// TIA Portal project "FABRICA DE TAPAS - TRANSPORTE -TUNEL DE ENFRIAMIENTO" (V17)

(* hardware
DEVICE "S7-1500/ET200MP station_1"  S7-1500 station
   slot 0: "Rail_0"  Rack  6ES7 590-1***0-0AA0
   slot 1: "CPU_PRINCIPAL"  CPU 1511-1 PN  6ES7 511-1AK02-0AB0  V2.8
      slot 3: "CPU display_1"  6ES7591-1AA00-0AA0
      slot 32768: "PROFINET interface_1"  X1
         slot 32769: "Port_1"  X1 P1
         slot 32770: "Port_2"  X1 P2
      slot 34817: "Virtual CP interface port_1"  Virtual CP interface port  Virtual CP interface port
DEVICE "HMI-TRANSPORTE"  KTP700 Basic PN
   slot 0: "HMI-TRANSPORTE"  KTP700 Basic PN  6AV2 123-2GB03-0AX0  17.0.0.0
   slot 1: "HMI_RT_1"  KTP700 Basic PN  6AV2 123-2GB03-0AX0  17.0.0.0
   slot 5: "HMI-TRANSPORTE.IE_CP_1"  PROFINET Interface  17.0.0.0
      slot 1: "PROFINET Interface_1"  PROFINET Interface
         slot 1: "Port_1"  Port
DEVICE "TUNEL-1"  KTP700 Basic PN
   slot 0: "TUNEL-1"  KTP700 Basic PN  6AV2 123-2GB03-0AX0  17.0.0.0
   slot 1: "HMI_RT_2"  KTP700 Basic PN  6AV2 123-2GB03-0AX0  17.0.0.0
   slot 5: "TUNEL-1.IE_CP_1"  PROFINET Interface  17.0.0.0
      slot 1: "PROFINET Interface_1"  PROFINET Interface
         slot 1: "Port_1"  Port
DEVICE "TUNEL-2"  KTP700 Basic PN
   slot 0: "TUNEL-2"  KTP700 Basic PN  6AV2 123-2GB03-0AX0  17.0.0.0
   slot 1: "HMI_RT_3"  KTP700 Basic PN  6AV2 123-2GB03-0AX0  17.0.0.0
   slot 5: "TUNEL-2.IE_CP_1"  PROFINET Interface  17.0.0.0
      slot 1: "PROFINET Interface_1"  PROFINET Interface
         slot 1: "Port_1"  Port
DEVICE "ET 200SP station_1"  ET 200SP-Station
   slot 0: "Rack_0"  Rack  6ES5 710-8MAx1
   slot 0: "TRANSPORTE"  IM 155-6 PN ST  6ES7 155-6AU01-0BN0  V4.2
   slot 1: "DI 16x24VDC ST_1"  DI 16x24VDC ST  6ES7 131-6BH01-0BA0  V0.0
      slot 1: "DI 16x24VDC ST_1"  DI 16x24VDC ST
   slot 2: "DQ 16x24VDC/0.5A ST_1"  DQ 16x24VDC/0.5A ST  6ES7 132-6BH01-0BA0  V0.0
      slot 1: "DQ 16x24VDC/0.5A ST_1"  DQ 16x24VDC/0.5A ST
   slot 3: "Server module_1"  Server module  6ES7 193-6PA00-0AA0  V1.1
      slot 1: "Server module_1"  Server module
   slot 127: "BA 2xRJ45"  BA 2xRJ45  6ES7 193-6AR00-0AA0  V0.0
      slot 1: "Port_1"  X1 P1 R  6ES7 193-6AR00-0AA0  V0.0
      slot 2: "Port_2"  X1 P2 R  6ES7 193-6AR00-0AA0  V0.0
DEVICE "ET 200SP station_2"  ET 200SP-Station
   slot 0: "Rack_0"  Rack  6ES5 710-8MAx1
   slot 0: "TUNEL_1"  IM 155-6 PN ST  6ES7 155-6AU01-0BN0  V4.2
   slot 1: "DI 16x24VDC ST_1"  DI 16x24VDC ST  6ES7 131-6BH01-0BA0  V0.0
      slot 1: "DI 16x24VDC ST_1"  DI 16x24VDC ST
   slot 2: "DQ 16x24VDC/0.5A ST_1"  DQ 16x24VDC/0.5A ST  6ES7 132-6BH01-0BA0  V0.0
      slot 1: "DQ 16x24VDC/0.5A ST_1"  DQ 16x24VDC/0.5A ST
   slot 3: "Server module_1"  Server module  6ES7 193-6PA00-0AA0  V1.1
      slot 1: "Server module_1"  Server module
   slot 127: "BA 2xRJ45"  BA 2xRJ45  6ES7 193-6AR00-0AA0  V0.0
      slot 1: "Port_1"  X1 P1 R  6ES7 193-6AR00-0AA0  V0.0
      slot 2: "Port_2"  X1 P2 R  6ES7 193-6AR00-0AA0  V0.0
DEVICE "ET 200SP station_3"  ET 200SP-Station
   slot 0: "Rack_0"  Rack  6ES5 710-8MAx1
   slot 0: "TUNEL_2"  IM 155-6 PN ST  6ES7 155-6AU01-0BN0  V4.2
   slot 1: "DI 16x24VDC ST_1"  DI 16x24VDC ST  6ES7 131-6BH01-0BA0  V0.0
      slot 1: "DI 16x24VDC ST_1"  DI 16x24VDC ST
   slot 2: "DQ 16x24VDC/0.5A ST_1"  DQ 16x24VDC/0.5A ST  6ES7 132-6BH01-0BA0  V0.0
      slot 1: "DQ 16x24VDC/0.5A ST_1"  DQ 16x24VDC/0.5A ST
   slot 3: "Server module_1"  Server module  6ES7 193-6PA00-0AA0  V1.1
      slot 1: "Server module_1"  Server module
   slot 127: "BA 2xRJ45"  BA 2xRJ45  6ES7 193-6AR00-0AA0  V0.0
      slot 1: "Port_1"  X1 P1 R  6ES7 193-6AR00-0AA0  V0.0
      slot 2: "Port_2"  X1 P2 R  6ES7 193-6AR00-0AA0  V0.0
*)

// ===== PLC "CPU_PRINCIPAL"  CPU 1511-1 PN =====

VAR_GLOBAL   // PLC tag table "Default tag table"
   "System_Byte" AT %MB1000 : Byte;
   "FirstScan" AT %M1000.0 : Bool;
   "DiagStatusUpdate" AT %M1000.1 : Bool;
   "AlwaysTRUE" AT %M1000.2 : Bool;
   "AlwaysFALSE" AT %M1000.3 : Bool;
   "Clock_Byte" AT %MB2000 : Byte;
   "Clock_10Hz" AT %M2000.0 : Bool;
   "Clock_5Hz" AT %M2000.1 : Bool;
   "Clock_2.5Hz" AT %M2000.2 : Bool;
   "Clock_2Hz" AT %M2000.3 : Bool;
   "Clock_1.25Hz" AT %M2000.4 : Bool;
   "Clock_1Hz" AT %M2000.5 : Bool;
   "Clock_0.625Hz" AT %M2000.6 : Bool;
   "Clock_0.5Hz" AT %M2000.7 : Bool;
   "Tag_1" AT %M3000.0 : Bool;
   "Tag_2" AT %M3000.1 : Bool;
   "Tag_3" AT %M3000.3 : Bool;
   "Tag_4" AT %M3001.0 : Bool;
END_VAR

VAR_GLOBAL   // PLC tag table "Entradas Digitales tunel 1"
   "Paro_Emergencia_Tunel_1" AT %I10.0 : Bool;   // Contacto NC fisico
   "Reset_Falla_Tunel_1" AT %I10.1 : Bool;   // Contacto NC fisico
   "Modo_Local_Tunel_1" AT %I10.2 : Bool;   // Contacto NO fisico
   "Modo_Automatico_Tunel_1" AT %I10.3 : Bool;   // Contacto NO fisico
   "Presostato_Tunel_1" AT %I10.4 : Bool;   // Contacto NO fisico
   "Confirmacion_banda_tunel_1" AT %I10.5 : Bool;   // Contacto NO de KM1 confirmacion arranque de banda
   "Confirmacion_aspirador_tunel_1" AT %I10.6 : Bool;   // Contacto NO de KM2 confirmacion arranque de aspirador
   "Confirmacion_Ventilador_tunel_1" AT %I10.7 : Bool;   // Contacto NO de KM2 confirmacion arranque de Ventilador
   "Confirmacion_Vibrador_tunel_1" AT %I11.0 : Bool;   // Contacto NO de KM2 confirmacion arranque de Vibracion
   "Señal_de_fallo_banda_tunel_1" AT %I11.1 : Bool;   // Contacto NO Guardamotor QM1
   "Señal_de_fallo_aspirador_tunel_1" AT %I11.2 : Bool;   // Contacto NO Guardamotor QM2
   "Señal_de_fallo_ventilador_tunel_1" AT %I11.3 : Bool;   // Contacto NO Guardamotor QM3
   "Señal_de_fallo_vibrador_tunel_1" AT %I11.4 : Bool;   // Contacto NO Guardamotor QM4
   "Confirmacion_trafico_tapas" AT %I11.5 : Bool;   // Señal de Plastificadora para indicar que hay tapas
   "Señal_Intercambio" AT %I11.6 : Bool;
   "Reserva" AT %I11.7 : Bool;
END_VAR

VAR_GLOBAL   // PLC tag table "Entradas Digitales Tunel 2"
   "Paro_Emergencia_Tunel_2" AT %I20.0 : Bool;   // Contacto NC fisico
   "Reset_Falla_Tunel_2" AT %I20.1 : Bool;   // Contacto NC fisico
   "Modo_Local_Tunel_2" AT %I20.2 : Bool;   // Contacto NO fisico
   "Modo_Automatico_Tunel_2" AT %I20.3 : Bool;   // Contacto NO fisico
   "Presostato_Tunel_2" AT %I20.4 : Bool;   // Contacto NO fisico
   "Confirmacion_banda_tunel_2" AT %I20.5 : Bool;   // Contacto NO de KM1 confirmacion arranque de banda
   "Confirmacion_aspirador_tunel_2" AT %I20.6 : Bool;   // Contacto NO de KM2 confirmacion arranque de aspirador
   "Confirmacion_Ventilador_tunel_2" AT %I20.7 : Bool;   // Contacto NO de KM2 confirmacion arranque de Ventilador
   "Confirmacion_Vibrador_tunel_2" AT %I21.0 : Bool;   // Contacto NO de KM2 confirmacion arranque de Vibracion
   "Señal_de_fallo_banda_tunel_2" AT %I21.1 : Bool;   // Contacto NO Guardamotor QM1
   "Señal_de_fallo_aspirador_tunel_2" AT %I21.2 : Bool;   // Contacto NO Guardamotor QM2
   "Señal_de_fallo_ventilador_tunel_2" AT %I21.3 : Bool;   // Contacto NO Guardamotor QM3
   "Señal_de_fallo_vibrador_tunel_2" AT %I21.4 : Bool;   // Contacto NO Guardamotor QM4
   "Confirmacion_trafico_tapas_2" AT %I21.5 : Bool;   // Señal de Plastificadora para indicar que hay tapas
   "Señal_Intercambio_2" AT %I21.6 : Bool;
   "Reserva_2" AT %I21.7 : Bool;
END_VAR

VAR_GLOBAL   // PLC tag table "Salidas Digitales Tunel 1"
   "Motor_banda_tunel_1" AT %Q10.0 : Bool;
   "Motor_aspirador_tunel_!" AT %Q10.1 : Bool;
   "Motor_ventilador_tunel_1" AT %Q10.2 : Bool;
   "Motor_vibrador_tunel_1" AT %Q10.3 : Bool;
   "Desviar_cajas_derecha_Tunel_1" AT %Q10.4 : Bool;
   "Desviar_cajas_izquierda_Tunel_1" AT %Q10.5 : Bool;
   "Valvula_soplado_Tunel_1" AT %Q10.6 : Bool;
   "Bajar_cuchara_Tunel_1" AT %Q10.7 : Bool;
   "Subir_Cuchara_Tunel_1" AT %Q11.0 : Bool;
   "Señalizacion_Roja_Tunel_1" AT %Q11.1 : Bool;
   "Señalizacion_azul_tunel_1" AT %Q11.2 : Bool;
   "Señalizacion_operacion_verde_tunel_1" AT %Q11.3 : Bool;
   "Reserva_1_tunel_1" AT %Q11.4 : Bool;
   "Señal_Intercambio_Tunel_1" AT %Q11.5 : Bool;
   "Reserva_2_tunel_1" AT %Q11.6 : Bool;
   "Reserva_3_tunel_1" AT %Q11.7 : Bool;
END_VAR

VAR_GLOBAL   // PLC tag table "Salidas Digitales Tunel 2"
   "Motor_banda_tunel_2" AT %Q20.0 : Bool;
   "Motor_aspirador_tunel_2" AT %Q20.1 : Bool;
   "Motor_ventilador_tunel_2" AT %Q20.2 : Bool;
   "Motor_vibrador_tunel_2" AT %Q20.3 : Bool;
   "Desviar_cajas_derecha_Tunel_2" AT %Q20.4 : Bool;
   "Desviar_cajas_izquierda_Tunel_2" AT %Q20.5 : Bool;
   "Valvula_soplado_Tunel_2" AT %Q20.6 : Bool;
   "Bajar_cuchara_Tunel_2" AT %Q20.7 : Bool;
   "Subir_Cuchara_Tunel_2" AT %Q21.0 : Bool;
   "Señalizacion_Roja_Tunel_2" AT %Q21.1 : Bool;
   "Señalizacion_Azul_tunel_2" AT %Q21.2 : Bool;
   "Señalizacion_operacion_Verde_tunel_2" AT %Q21.3 : Bool;
   "Reserva_1_tunel_2" AT %Q21.4 : Bool;
   "Señal_Intercambio_Tunel_2" AT %Q21.5 : Bool;
   "Reserva_2_tunel_2" AT %Q21.6 : Bool;
   "Reserva_3_tunel_2" AT %Q21.7 : Bool;
END_VAR

VAR_GLOBAL   // PLC tag table "Entradas Digitales Transporte"
   "Paro de emergencia transporte" AT %I0.0 : Bool;   // SEÑAL NC
   "Reset Falla transporte" AT %I0.1 : Bool;   // SEÑAL NC
   "Orden Llenado Tolva 1" AT %I0.2 : Bool;
   "Orden Llenado Tolva 2" AT %I0.3 : Bool;
   "Presostato" AT %I0.4 : Bool;
   "Sensor_Nivel_Tolva_Reserva" AT %I0.5 : Bool;
   "Sensor_Nivel_Tolva_Tunel_1" AT %I0.6 : Bool;
   "Sensor_Nivel_Tolva_Tunel_2" AT %I0.7 : Bool;
   "Tolva_descarga_Tolva" AT %I1.0 : Bool;
   "Señal Retorno QM1" AT %I1.1 : Bool;
   "Señal Retorno QM2" AT %I1.2 : Bool;
   "Señal Retorno QM3" AT %I1.3 : Bool;
   "Señal Retorno QM4" AT %I1.4 : Bool;
   "Señal PILZ" AT %I1.5 : Bool;
   "Automatico" AT %I1.6 : Bool;
   "Manual" AT %I1.7 : Bool;
END_VAR

VAR_GLOBAL   // PLC tag table "Salidas Digitales Transporte"
   "M1 (motor elevador)" AT %Q0.0 : Bool;
   "M2 (motor traslado)" AT %Q0.1 : Bool;
   "M3 (motor llenado tolvas)" AT %Q0.2 : Bool;
   "KM4 (motor entrada tolvas suministro)" AT %Q0.3 : Bool;
   "YV1  (Restriccion paso)" AT %Q0.4 : Bool;
   "YV2 (compuertas)" AT %Q0.5 : Bool;
   "YV3 (Electrovalvula paso tolva 1)" AT %Q0.6 : Bool;
   "YV2A (electrovalvula paso tolva 2)" AT %Q0.7 : Bool;
   "Vibrador" AT %Q1.0 : Bool;
   "Piloto de falla color rojo" AT %Q1.1 : Bool;
   "Piloto de paro programado color azul" AT %Q1.2 : Bool;
   "piloto de encendido ok color verde" AT %Q1.3 : Bool;
   "Reserva 1" AT %Q1.4 : Bool;
   "Reserva 2" AT %Q1.5 : Bool;
   "Reserva 3" AT %Q1.6 : Bool;
   "Reserva 4" AT %Q1.7 : Bool;
END_VAR

VAR_GLOBAL   // PLC tag table "CONSIGNAS_TEMPORIZADORES"
   "TEMPORIZADOR_PASO_TAPAS_TUNEL_1" AT %MW0 : Int;
   "TEMPORIZADOR_BLOQUEO_TAPAS_TUNEL_1" AT %MW2 : Int;
   "TEMPORIZADOR_CAMBIO_DE_LLENADO_CAJA_TUNEL_1" AT %MW4 : Int;
   "TEMPORIZADOR_PASO_TAPAS_TUNEL_2" AT %MW6 : Int;
   "TEMPORIZADOR_BLOQUEO_TAPAS_TUNEL_2" AT %MW8 : Int;
   "TEMPORIZADOR_CAMBIO_DE_LLENADO_CAJA_TUNEL_2" AT %MW10 : Int;
END_VAR

DATA_BLOCK "BOTONERA_HMI_TUNEL_1"   // DB1
{ S7_Optimized_Access := 'TRUE' }
VERSION : 0.1
   VAR
      KM1_INICIO_MANUAL_BANDA_TUNEL_1 : Bool;
      KM1_STOP_MANUAL_BANDA_TUNEL_1 : Bool;
      KM2_INICIO_MANUAL_ASPIRADOR_TUNEL_1 : Bool;
      KM2_STOP_MANUAL_ASPIRADOR_TUNEL_1 : Bool;
      KM3_INICIO_MANUAL_VENTILADOR_TUNEL_1 : Bool;
      KM3_STOP_MANUAL_VENTILADOR_TUNEL_1 : Bool;
      KM4_INICIO_MANUAL_VIBRADOR_TUNEL_1 : Bool;
      KM4_STOP_MANUAL_VIBRADOR_TUNEL_1 : Bool;
      SUBIR_CUCHARA_TUNEL_1 : Bool;
      BAJAR_CUCHARA_TUNEL_1 : Bool;
      CARGADOR_CAJAS_DERECHA_TUNEL_1 : Bool;
      CARGADOR_CAJAS_IZQUIERDA_TUNEL_1 : Bool;
   END_VAR
BEGIN
END_DATA_BLOCK

DATA_BLOCK "BOTONERA_HMI_TUNEL_2"   // DB2
{ S7_Optimized_Access := 'TRUE' }
VERSION : 0.1
   VAR
      KM1_INICIO_MANUAL_BANDA_TUNEL_2 : Bool;
      KM1_STOP_MANUAL_BANDA_TUNEL_2 : Bool;
      KM2_INICIO_MANUAL_ASPIRADOR_TUNEL_2 : Bool;
      KM2_STOP_MANUAL_ASPIRADOR_TUNEL_2 : Bool;
      KM3_INICIO_MANUAL_VENTILADOR_TUNEL_2 : Bool;
      KM3_STOP_MANUAL_VENTILADOR_TUNEL_2 : Bool;
      KM4_INICIO_MANUAL_VIBRADOR_TUNEL_2 : Bool;
      KM4_STOP_MANUAL_VIBRADOR_TUNEL_2 : Bool;
      SUBIR_CUCHARA_TUNEL_2 : Bool;
      BAJAR_CUCHARA_TUNEL_2 : Bool;
      CARGADOR_CAJAS_DERECHA_TUNEL_2 : Bool;
      CARGADOR_CAJAS_IZQUIERDA_TUNEL_2 : Bool;
   END_VAR
BEGIN
END_DATA_BLOCK

DATA_BLOCK "BOTONERA_HMI_TRANSPORTE"   // DB3
{ S7_Optimized_Access := 'TRUE' }
VERSION : 0.1
   VAR
      KM1_INICIO_MANUAL_ELEVADOR_TRANSPORTE : Bool;
      KM1_STOP_MANUAL_ELEVADOR_TRANSPORTE : Bool;
      KM2_INICIO_MANUAL_TRANSPORTE_GENERAL_TRANSPORTE : Bool;
      KM2_STOP_MANUAL_TRANSPORTE_GENERAL_TRANSPORTE : Bool;
      KM3_INICIO_MANUAL_TOLVAS_TRANSPORTE : Bool;
      KM3_STOP_MANUAL_TOLVAS_TRANSPORTE : Bool;
      "KM4_ INICIO_MANUAL_VIBRADOR_TRANSPORTE" : Bool;
      KM4_STOP_MANUAL_VIBRADOR_TRANSPORTE : Bool;
      "DESVIADOR_DE BANDA_NEUMATICO_ACTIVAR_MANUAL" : Bool;
      "DESVIADOR_DE BANDA_NEUMATICO_DESACTIVAR_MANUAL" : Bool;
      COMPUERTA_TOLVA_RESERVA_NEUMATICO_ACTIVAR_MANUAL : Bool;
      COMPUERTA_TOLVA_RESERVA_NEUMATICO_DESACTIVAR_MANUAL : Bool;
      LLENADO_TOLVAS_ACTIVAR_MANUAL : Bool;
      LLENADO_TOLVAS_DESACTIVAR_MANUAL : Bool;
   END_VAR
BEGIN
END_DATA_BLOCK

DATA_BLOCK "PERMISOS_DE_MARCHA_TUNEL_1"   // DB4
{ S7_Optimized_Access := 'TRUE' }
VERSION : 0.1
   VAR
      BANDA_TUNEL_1_AUTOMATICO : Bool;
      BANDA_TUNEL_1_MANUAL : Bool;
      ASPIRADOR_TUNEL_1_AUTOMATICO : Bool;
      ASPIRADOR_TUNEL_1_MANUAL : Bool;
      VENTILADOR_TUNEL_1_AUTOMATICO : Bool;
      VENTILADOR_TUNEL_1_MANUAL : Bool;
      VIBRADOR_TUNEL_1_AUTOMATICO : Bool;
      VIBRADOR_TUNEL_1_MANUAL : Bool;
      ABRIR_CUCHARA_TUNEL_1_AUTOMATICO : Bool;
      CERRAR_CUCHARA_TUNEL_1_AUTOMATICO : Bool;
      CERRAR_CUCHARA_TUNEL_1_MANUAL : Bool;
      ABRIR_CUCHARA_TUNEL_1_MANUAL : Bool;
      CAJA_DERECHA_TUNEL_1_AUTOMATICO : Bool;
      CAJA_DERECHA_TUNEL_1_MANUAL : Bool;
      CAJA_IZQUIERDA_TUNEL_1_AUTOMATICO : Bool;
      CAJA_IZQUIERDA_TUNEL_1_MANUAL : Bool;
   END_VAR
BEGIN
END_DATA_BLOCK

DATA_BLOCK "PERMISOS_DE_MARCHA_TUNEL_2"   // DB5
{ S7_Optimized_Access := 'TRUE' }
VERSION : 0.1
   VAR
      BANDA_TUNEL_2_AUTOMATICO : Bool;
      BANDA_TUNEL_2_MANUAL : Bool;
      ASPIRADOR_TUNEL_2_AUTOMATICO : Bool;
      ASPIRADOR_TUNEL_2_MANUAL : Bool;
      VENTILADOR_TUNEL_2_AUTOMATICO : Bool;
      VENTILADOR_TUNEL_2_MANUAL : Bool;
      VIBRADOR_TUNEL_2_AUTOMATICO : Bool;
      VIBRADOR_TUNEL_2_MANUAL : Bool;
      ABRIR_CUCHARA_TUNEL_2_AUTOMATICO : Bool;
      CERRAR_CUCHARA_TUNEL_2_MANUAL : Bool;
      CERRAR_CUCHARA_TUNEL_2_AUTOMATICO : Bool;
      ABRIR_CUCHARA_TUNEL_2_MANUAL : Bool;
      CAJA_DERECHA_TUNEL_2_AUTOMATICO : Bool;
      CAJA_DERECHA_TUNEL_2_MANUAL : Bool;
      CAJA_IZQUIERDA_TUNEL_2_AUTOMATICO : Bool;
      CAJA_IZQUIERDA_TUNEL_2_MANUAL : Bool;
   END_VAR
BEGIN
END_DATA_BLOCK

DATA_BLOCK "PERMISOS_GENERALES"   // DB6
{ S7_Optimized_Access := 'TRUE' }
VERSION : 0.1
   VAR
      TUNEL_1_DESHABILITADO : Bool;
      TUNEL_2_DESHABILITADO : Bool;
      MODO_LOCAL_2 : Bool;
      MODO_AUTOMATICO_2 : Bool;
      MODO_AUTOMATICO_1 : Bool;
      MODO_LOCAL_1 : Bool;
      MODO_AUTOMATICO_TRANSPORTE : Bool;
      MODO_MANUAL_TRANSPORTE : Bool;
      TRANSPORTE_DESHABILITADO : Bool;
   END_VAR
BEGIN
END_DATA_BLOCK

DATA_BLOCK "MEMORIAS_DE_ESTADOS_TUNEL_1"   // DB7
{ S7_Optimized_Access := 'TRUE' }
VERSION : 0.1
   VAR
      CAMBIO_ESTADO_AUTOMATICO_TUNEL_1 : Bool;
      CAMBIO_ESTADO_MANUAL_TUNEL_1 : Bool;
      TRANSICION_CAJA_TUNEL_FLANCO : Bool;
      TRANSICION_CAJA_TUNEL_1 : Bool;
      INICIO_CONTEO_CAMBIO_CAJA_TUNEL_1 : Bool;
      CUENTA_11K_TAPAS : Bool;
      CONTEO_TAPAS_TUNEL_1 : Bool;
      CAMBIO_ESTADO_TUNEL_1_PRESENTE : Bool;
   END_VAR
BEGIN
END_DATA_BLOCK

DATA_BLOCK "TIEMPOS_TUNEL_1"   // DB9
{ S7_Optimized_Access := 'TRUE' }
VERSION : 0.1
   VAR
      PASO_TAPAS_TUNEL_1 : Int;
      BLOQUEO_TAPAS_TUNEL_1 : Int;
      CAMBIO_CAJA_TUNEL_1 : Int;
      TIEMPO_TOTAL_PASO_BLOQUEO : Int;
   END_VAR
BEGIN
END_DATA_BLOCK

DATA_BLOCK "MEMORIAS_DE_ESTADOS_TUNEL_2"   // DB11
{ S7_Optimized_Access := 'TRUE' }
VERSION : 0.1
   VAR
      CAMBIO_ESTADO_AUTOMATICO_TUNEL_2 : Bool;
      CAMBIO_ESTADO_MANUAL_TUNEL_2 : Bool;
      TRANSICION_CAJA_TUNEL2_FLANCO : Bool;
      TRANSICION_CAJA_TUNEL_2 : Bool;
      INICIO_CONTEO_CAMBIO_CAJA_TUNEL_2 : Bool;
      CUENTA_11K_TAPAS_2 : Bool;
      CONTEO_TAPAS_TUNEL_2 : Bool;
      CAMBIO_ESTADO_TUNEL_2_PRESENTE : Bool;
   END_VAR
BEGIN
END_DATA_BLOCK

DATA_BLOCK "TIEMPOS_TUNEL_2"   // DB13
{ S7_Optimized_Access := 'TRUE' }
VERSION : 0.1
   VAR
      PASO_TAPAS_TUNEL_2 : Int;
      BLOQUEO_TAPAS_TUNEL_2 : Int;
      CAMBIO_CAJA_TUNEL_2 : Int;
      TIEMPO_TOTAL2_PASO_BLOQUEO : Int;
   END_VAR
BEGIN
END_DATA_BLOCK

DATA_BLOCK "MEMORIAS_DE_ESTADO_TRANSPORTE"   // DB15
{ S7_Optimized_Access := 'TRUE' }
VERSION : 0.1
   VAR
      CAMBIO_DE_ESTADO_PRESENTA : Bool;
      "TRANSICION A MANUAL" : Bool;
      "TRANSICION A AUTOMATICO" : Bool;
   END_VAR
BEGIN
END_DATA_BLOCK

DATA_BLOCK "PERMISOS_DE_MARCHA_TRANSPORTE"   // DB16
{ S7_Optimized_Access := 'TRUE' }
VERSION : 0.1
   VAR
      ELEVADOR_MANUAL : Bool;
      ELEVADOR_AUTOMATICO : Bool;
      CIRCULACION_MANUAL : Bool;
      CIRCULACION_AUTOMATICO : Bool;
      TOLVA_RESERVA_MANUAL : Bool;
      TOLVA_RESERVA_AUTOMATICO : Bool;
      VIBRADOR_MANUAL : Bool;
      VIBRADOR_AUTOMATICO : Bool;
      ELECTROVALVULA_RESTRICCION_PASO_MANUAL : Bool;
      ELECTROVALVULA_RESTRICCION_PASO_AUTOMATICO : Bool;
      ELECTROVALVULA_COMPUERTA_TOLVA_RESERVA_MANUAL : Bool;
      ELECTROVALVULA_COMPUERTA_TOLVA_RESERVA_AUTOMATICO : Bool;
      ELECTROVALVULA_LLENADO_TOLVA_1_MANUAL : Bool;
      ELECTROVALVULA_LLENADO_TOLVA_1_AUTOMATICO : Bool;
      ELECTROVALVULA_LLENADO_TOLVA_2_MANUAL : Bool;
      MOTOR_LLENADO_TOLVAS_MANUAL : Bool;
      MOTOR_LLENADO_TOLVAS_AUTOMATICO : Bool;
      ELECTROVALVULA_LLENADO_TOLVA_2_AUTOMATICO : Bool;
   END_VAR
BEGIN
END_DATA_BLOCK

DATA_BLOCK "FALLAS_TUNEL_1"   // DB17
{ S7_Optimized_Access := 'TRUE' }
VERSION : 0.1
   VAR
      MOTOR_AVERIADO_TUNEL_1 : Bool;
      PRESOSTATO_OFF_TUNEL_1 : Bool;
      PARADA_EMERGENCIA_TUNEL_1 : Bool;
      EQUIPO_OPERANDO_EN_AUTOMATICO_TUNEL_1 : Bool;
      NO_TAPAS_TUNEL_1 : Bool;
      EQUIPO_OPERANDO_EN_MANUAL_TUNEL_1 : Bool;
   END_VAR
BEGIN
END_DATA_BLOCK

DATA_BLOCK "FALLAS_TUNEL_2"   // DB18
{ S7_Optimized_Access := 'TRUE' }
VERSION : 0.1
   VAR
      MOTOR_AVERIADO_TUNEL_2 : Bool;
      PRESOSTATO_OFF_TUNEL_2 : Bool;
      PARADA_EMERGENCIA_TUNEL_2 : Bool;
      EQUIPO_OPERANDO_EN_AUTOMATICO_TUNEL_2 : Bool;
      NO_TAPAS_TUNEL_2 : Bool;
      EQUIPO_OPERANDO_EN_MANUAL_TUNEL_2 : Bool;
   END_VAR
BEGIN
END_DATA_BLOCK

DATA_BLOCK "ANIMACIONES"   // DB19
{ S7_Optimized_Access := 'TRUE' }
VERSION : 0.1
   VAR
      MOVIMIENTO_FLECHA_TUNEL_2 : Int;
      MOVIMIENTO_FLECHA_VIBRADOR_TUNEL_2 : Int;
      MOVIMIENTO_FLECHA_VIBRADOR_TUNEL_1 : Int;
      MOVIMIENTO_FLECHA_BANDA_TUNEL_1 : Int;
      BANDA_1_ENCENDIDA : Bool;
      BANDA_2_ENCENDIDA : Bool;
   END_VAR
BEGIN
END_DATA_BLOCK

DATA_BLOCK "Alarmas_tunel_1"   // DB24
{ S7_Optimized_Access := 'FALSE' }
VERSION : 0.1
   VAR
      "BANDA EN FALLA" : Bool;
      "ASPIRADOR EN FALLA" : Bool;
      "VENTILADOR EN FALLA" : Bool;
      "VIBRADOR EN FALLA" : Bool;
      "PRESOSTATO OFF" : Bool;
      "SIN SUMINISTRO TAPAS" : Bool;
      "PARO DE EMERGENCIA" : Bool;
   END_VAR
BEGIN
END_DATA_BLOCK

// folder: System blocks/Program resources

DATA_BLOCK "TIEMPO_GENERAL_TUNEL_1"   // DB8
{ S7_Optimized_Access := 'TRUE' }
AUTHOR : Simatic
FAMILY : IEC
NAME : CNTR
VERSION : 1.0
// stored: InstanceOfName IEC_COUNTER
"IEC_COUNTER"
BEGIN
END_DATA_BLOCK

DATA_BLOCK "CONTADOR_CAMBIO_CAJA_TUNEL_1"   // DB10
{ S7_Optimized_Access := 'TRUE' }
AUTHOR : Simatic
FAMILY : IEC
NAME : CNTR
VERSION : 1.0
// stored: InstanceOfName IEC_COUNTER
"IEC_COUNTER"
BEGIN
END_DATA_BLOCK

DATA_BLOCK "TIEMPO_GENERAL_TUNEL_2"   // DB12
{ S7_Optimized_Access := 'TRUE' }
AUTHOR : Simatic
FAMILY : IEC
NAME : CNTR
VERSION : 1.0
// stored: InstanceOfName IEC_COUNTER
"IEC_COUNTER"
BEGIN
END_DATA_BLOCK

DATA_BLOCK "CONTADOR_CAMBIO_CAJA_TUNEL_2"   // DB14
{ S7_Optimized_Access := 'TRUE' }
AUTHOR : Simatic
FAMILY : IEC
NAME : CNTR
VERSION : 1.0
// stored: InstanceOfName IEC_COUNTER
"IEC_COUNTER"
BEGIN
END_DATA_BLOCK

DATA_BLOCK "AVANCE_FLECHA_TUNEL_1"   // DB20
{ S7_Optimized_Access := 'TRUE' }
AUTHOR : Simatic
FAMILY : IEC
NAME : CNTR
VERSION : 1.0
// stored: InstanceOfName IEC_COUNTER
"IEC_COUNTER"
BEGIN
END_DATA_BLOCK

DATA_BLOCK "AVANCE_FLECHA_TUNEL_2"   // DB21
{ S7_Optimized_Access := 'TRUE' }
AUTHOR : Simatic
FAMILY : IEC
NAME : CNTR
VERSION : 1.0
// stored: InstanceOfName IEC_COUNTER
"IEC_COUNTER"
BEGIN
END_DATA_BLOCK

DATA_BLOCK "VIBRADOR_FLECHA_TUNEL_1"   // DB22
{ S7_Optimized_Access := 'TRUE' }
AUTHOR : Simatic
FAMILY : IEC
NAME : CNTR
VERSION : 1.0
// stored: InstanceOfName IEC_COUNTER
"IEC_COUNTER"
BEGIN
END_DATA_BLOCK

DATA_BLOCK "VIBRADOR_FLECHA_TUNEL_2"   // DB23
{ S7_Optimized_Access := 'TRUE' }
AUTHOR : Simatic
FAMILY : IEC
NAME : CNTR
VERSION : 1.0
// stored: InstanceOfName IEC_COUNTER
"IEC_COUNTER"
BEGIN
END_DATA_BLOCK

// folder: (top level)

FUNCTION "MODO_REMOTO_TUNEL_1" : Void   // FC1, LAD
{ S7_Optimized_Access := 'TRUE' }
VERSION : 0.1
   VAR_TEMP   // added for the SCL form of the ladder/FBD networks
      _w1 : Bool;
      _w2 : Bool;
      _w3 : Bool;
      _w4 : Bool;
   END_VAR
BEGIN

REGION Network 1
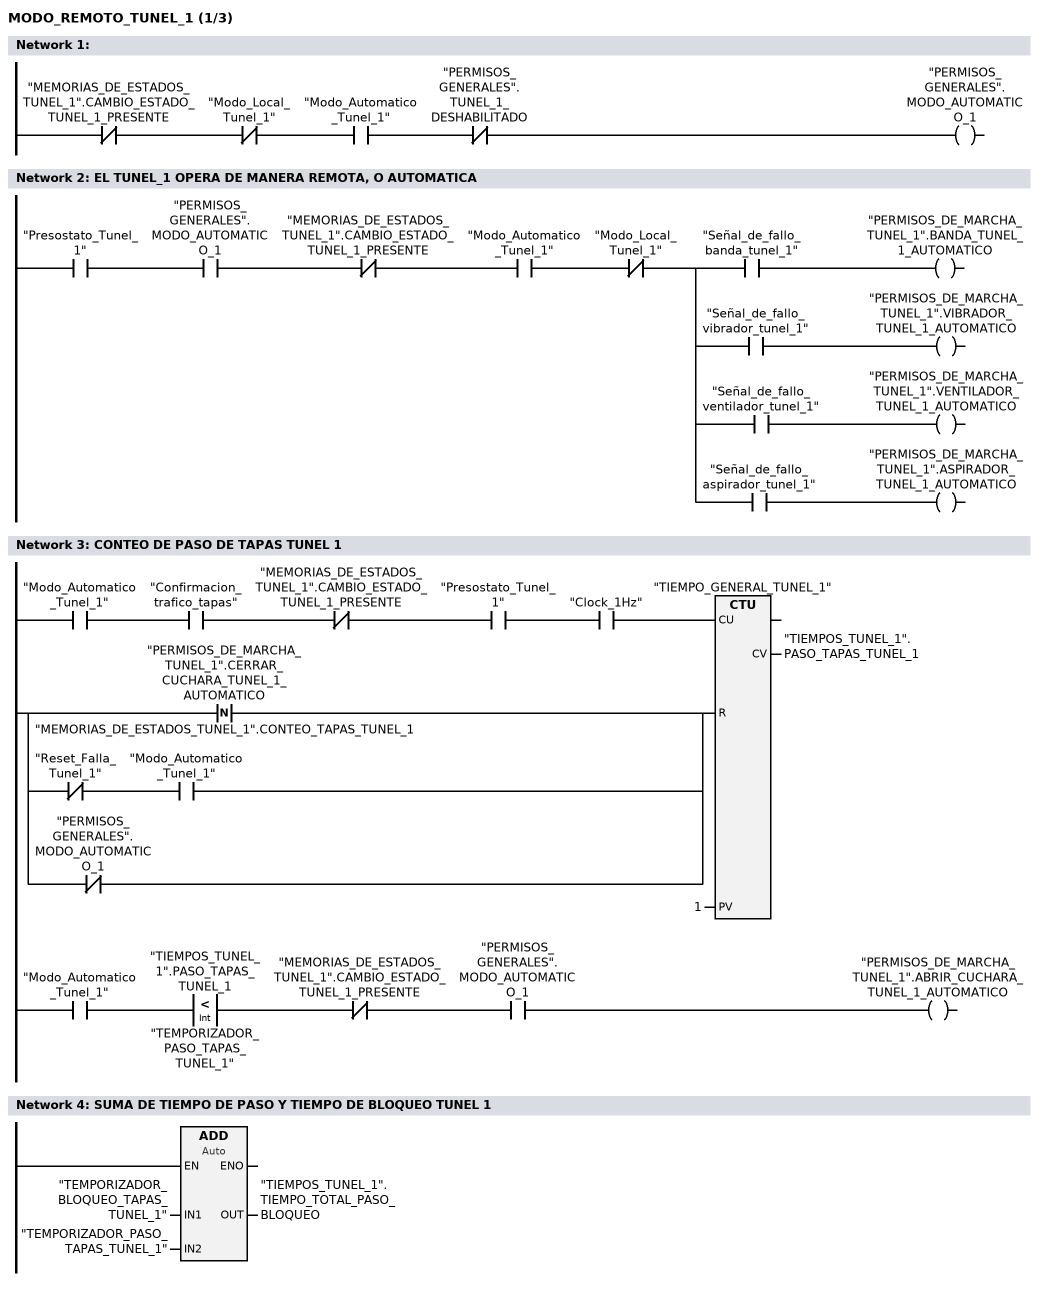
   RUNG wire#powerrail
      I_Contact( "MEMORIAS_DE_ESTADOS_TUNEL_1".CAMBIO_ESTADO_TUNEL_1_PRESENTE )
      I_Contact( "Modo_Local_Tunel_1" )
      Contact( "Modo_Automatico_Tunel_1" )
      I_Contact( "PERMISOS_GENERALES".TUNEL_1_DESHABILITADO )
      Coil( "PERMISOS_GENERALES".MODO_AUTOMATICO_1 )
   END_RUNG
   // the same network as SCL:
   "PERMISOS_GENERALES".MODO_AUTOMATICO_1 := NOT "MEMORIAS_DE_ESTADOS_TUNEL_1".CAMBIO_ESTADO_TUNEL_1_PRESENTE AND NOT "Modo_Local_Tunel_1" AND "Modo_Automatico_Tunel_1" AND NOT "PERMISOS_GENERALES".TUNEL_1_DESHABILITADO;
END_REGION

REGION Network 2: EL TUNEL_1 OPERA DE MANERA REMOTA, O AUTOMATICA
   RUNG wire#powerrail
      Contact( "Presostato_Tunel_1" )
      Contact( "PERMISOS_GENERALES".MODO_AUTOMATICO_1 )
      I_Contact( "MEMORIAS_DE_ESTADOS_TUNEL_1".CAMBIO_ESTADO_TUNEL_1_PRESENTE )
      Contact( "Modo_Automatico_Tunel_1" )
      I_Contact( "Modo_Local_Tunel_1" )
      wire#w1
      Contact( "Señal_de_fallo_banda_tunel_1" )
      Coil( "PERMISOS_DE_MARCHA_TUNEL_1".BANDA_TUNEL_1_AUTOMATICO )
   END_RUNG
   RUNG wire#w1
      Contact( "Señal_de_fallo_vibrador_tunel_1" )
      Coil( "PERMISOS_DE_MARCHA_TUNEL_1".VIBRADOR_TUNEL_1_AUTOMATICO )
   END_RUNG
   RUNG wire#w1
      Contact( "Señal_de_fallo_ventilador_tunel_1" )
      Coil( "PERMISOS_DE_MARCHA_TUNEL_1".VENTILADOR_TUNEL_1_AUTOMATICO )
   END_RUNG
   RUNG wire#w1
      Contact( "Señal_de_fallo_aspirador_tunel_1" )
      Coil( "PERMISOS_DE_MARCHA_TUNEL_1".ASPIRADOR_TUNEL_1_AUTOMATICO )
   END_RUNG
   // the same network as SCL:
   #_w1 := "Presostato_Tunel_1" AND "PERMISOS_GENERALES".MODO_AUTOMATICO_1 AND NOT "MEMORIAS_DE_ESTADOS_TUNEL_1".CAMBIO_ESTADO_TUNEL_1_PRESENTE AND "Modo_Automatico_Tunel_1" AND NOT "Modo_Local_Tunel_1";
   "PERMISOS_DE_MARCHA_TUNEL_1".BANDA_TUNEL_1_AUTOMATICO := #_w1 AND "Señal_de_fallo_banda_tunel_1";
   "PERMISOS_DE_MARCHA_TUNEL_1".VIBRADOR_TUNEL_1_AUTOMATICO := #_w1 AND "Señal_de_fallo_vibrador_tunel_1";
   "PERMISOS_DE_MARCHA_TUNEL_1".VENTILADOR_TUNEL_1_AUTOMATICO := #_w1 AND "Señal_de_fallo_ventilador_tunel_1";
   "PERMISOS_DE_MARCHA_TUNEL_1".ASPIRADOR_TUNEL_1_AUTOMATICO := #_w1 AND "Señal_de_fallo_aspirador_tunel_1";
END_REGION

REGION Network 3: CONTEO DE PASO DE TAPAS TUNEL 1
   #_w1 := NOT "PERMISOS_DE_MARCHA_TUNEL_1".CERRAR_CUCHARA_TUNEL_1_AUTOMATICO AND "MEMORIAS_DE_ESTADOS_TUNEL_1".CONTEO_TAPAS_TUNEL_1;   // falling edge of "PERMISOS_DE_MARCHA_TUNEL_1".CERRAR_CUCHARA_TUNEL_1_AUTOMATICO
   "MEMORIAS_DE_ESTADOS_TUNEL_1".CONTEO_TAPAS_TUNEL_1 := "PERMISOS_DE_MARCHA_TUNEL_1".CERRAR_CUCHARA_TUNEL_1_AUTOMATICO;
   "TIEMPO_GENERAL_TUNEL_1".CTU(CU := "Modo_Automatico_Tunel_1" AND "Confirmacion_trafico_tapas" AND NOT "MEMORIAS_DE_ESTADOS_TUNEL_1".CAMBIO_ESTADO_TUNEL_1_PRESENTE AND "Presostato_Tunel_1" AND "Clock_1Hz",
                           R := #_w1 OR (NOT "Reset_Falla_Tunel_1" AND "Modo_Automatico_Tunel_1") OR NOT "PERMISOS_GENERALES".MODO_AUTOMATICO_1,
                           PV := 1,
                           CV => "TIEMPOS_TUNEL_1".PASO_TAPAS_TUNEL_1);
   "PERMISOS_DE_MARCHA_TUNEL_1".ABRIR_CUCHARA_TUNEL_1_AUTOMATICO := "Modo_Automatico_Tunel_1" AND ("TIEMPOS_TUNEL_1".PASO_TAPAS_TUNEL_1 < "TEMPORIZADOR_PASO_TAPAS_TUNEL_1") AND NOT "MEMORIAS_DE_ESTADOS_TUNEL_1".CAMBIO_ESTADO_TUNEL_1_PRESENTE AND "PERMISOS_GENERALES".MODO_AUTOMATICO_1;
END_REGION

REGION Network 4: SUMA DE TIEMPO DE PASO Y TIEMPO DE BLOQUEO TUNEL 1
   RUNG wire#powerrail
      Add(in1 := "TEMPORIZADOR_BLOQUEO_TAPAS_TUNEL_1", in2 := "TEMPORIZADOR_PASO_TAPAS_TUNEL_1", out => "TIEMPOS_TUNEL_1".TIEMPO_TOTAL_PASO_BLOQUEO)
   END_RUNG
   // the same network as SCL:
   "TIEMPOS_TUNEL_1".TIEMPO_TOTAL_PASO_BLOQUEO := "TEMPORIZADOR_BLOQUEO_TAPAS_TUNEL_1" + "TEMPORIZADOR_PASO_TAPAS_TUNEL_1";
END_REGION

REGION Network 5: CIERRE DE CUCHARRA PARA BLOQUEO DE TAPAS TUNEL 1
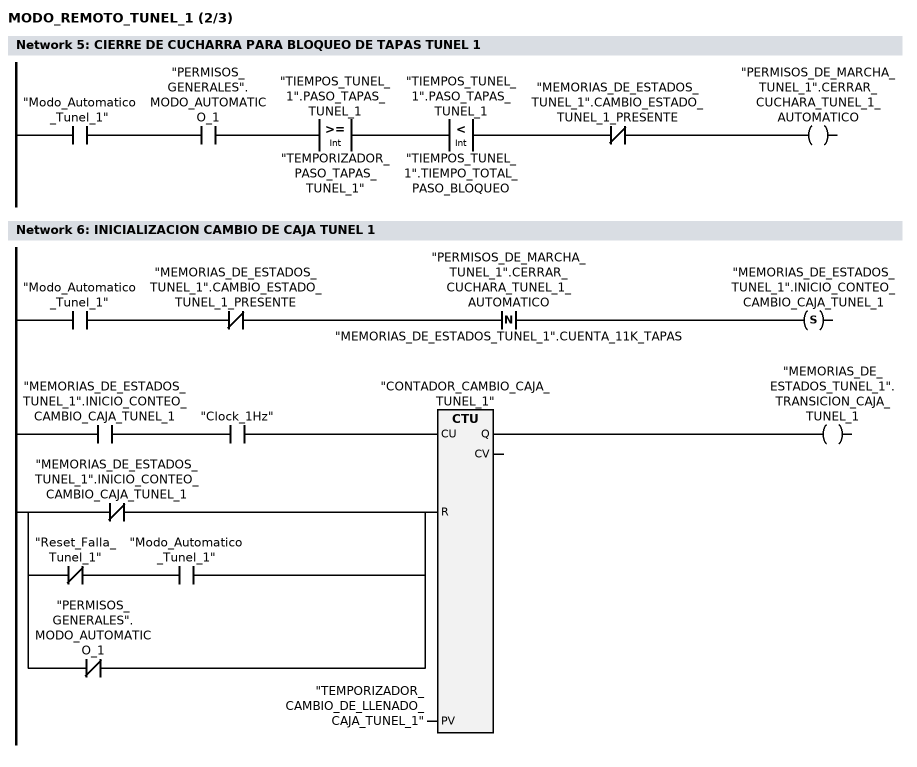
   RUNG wire#powerrail
      Contact( "Modo_Automatico_Tunel_1" )
      Contact( "PERMISOS_GENERALES".MODO_AUTOMATICO_1 )
      { S7_Templates := "SrcType := Int" } GE_Contact(in1 := "TIEMPOS_TUNEL_1".PASO_TAPAS_TUNEL_1, in2 := "TEMPORIZADOR_PASO_TAPAS_TUNEL_1")
      { S7_Templates := "SrcType := Int" } LT_Contact(in1 := "TIEMPOS_TUNEL_1".PASO_TAPAS_TUNEL_1, in2 := "TIEMPOS_TUNEL_1".TIEMPO_TOTAL_PASO_BLOQUEO)
      I_Contact( "MEMORIAS_DE_ESTADOS_TUNEL_1".CAMBIO_ESTADO_TUNEL_1_PRESENTE )
      Coil( "PERMISOS_DE_MARCHA_TUNEL_1".CERRAR_CUCHARA_TUNEL_1_AUTOMATICO )
   END_RUNG
   // the same network as SCL:
   "PERMISOS_DE_MARCHA_TUNEL_1".CERRAR_CUCHARA_TUNEL_1_AUTOMATICO := "Modo_Automatico_Tunel_1" AND "PERMISOS_GENERALES".MODO_AUTOMATICO_1 AND ("TIEMPOS_TUNEL_1".PASO_TAPAS_TUNEL_1 >= "TEMPORIZADOR_PASO_TAPAS_TUNEL_1") AND ("TIEMPOS_TUNEL_1".PASO_TAPAS_TUNEL_1 < "TIEMPOS_TUNEL_1".TIEMPO_TOTAL_PASO_BLOQUEO) AND NOT "MEMORIAS_DE_ESTADOS_TUNEL_1".CAMBIO_ESTADO_TUNEL_1_PRESENTE;
END_REGION

REGION Network 6: INICIALIZACION CAMBIO DE CAJA TUNEL 1
   #_w1 := "Modo_Automatico_Tunel_1" AND NOT "MEMORIAS_DE_ESTADOS_TUNEL_1".CAMBIO_ESTADO_TUNEL_1_PRESENTE AND NOT "PERMISOS_DE_MARCHA_TUNEL_1".CERRAR_CUCHARA_TUNEL_1_AUTOMATICO AND "MEMORIAS_DE_ESTADOS_TUNEL_1".CUENTA_11K_TAPAS;   // falling edge of "PERMISOS_DE_MARCHA_TUNEL_1".CERRAR_CUCHARA_TUNEL_1_AUTOMATICO
   "MEMORIAS_DE_ESTADOS_TUNEL_1".CUENTA_11K_TAPAS := "PERMISOS_DE_MARCHA_TUNEL_1".CERRAR_CUCHARA_TUNEL_1_AUTOMATICO;
   IF #_w1 THEN "MEMORIAS_DE_ESTADOS_TUNEL_1".INICIO_CONTEO_CAMBIO_CAJA_TUNEL_1 := TRUE; END_IF;
   "CONTADOR_CAMBIO_CAJA_TUNEL_1".CTU(CU := "MEMORIAS_DE_ESTADOS_TUNEL_1".INICIO_CONTEO_CAMBIO_CAJA_TUNEL_1 AND "Clock_1Hz",
                           R := NOT "MEMORIAS_DE_ESTADOS_TUNEL_1".INICIO_CONTEO_CAMBIO_CAJA_TUNEL_1 OR (NOT "Reset_Falla_Tunel_1" AND "Modo_Automatico_Tunel_1") OR NOT "PERMISOS_GENERALES".MODO_AUTOMATICO_1,
                           PV := "TEMPORIZADOR_CAMBIO_DE_LLENADO_CAJA_TUNEL_1");
   "MEMORIAS_DE_ESTADOS_TUNEL_1".TRANSICION_CAJA_TUNEL_1 := "CONTADOR_CAMBIO_CAJA_TUNEL_1".Q;
END_REGION

REGION Network 7: LOGICA DE CAMBIO DE CAJA TUNEL 1